
               Strg_TO_Chars(Strg:= CONCAT_STRING(IN1 := #TMP_strDef ,IN2 := DINT_TO_STRING(#INO_tDefects.tDefectsForReport.rgtDefects[#TMP_dIndexDef].dCoreWidth_um)),
                         pChars:=#TMP_dIndex,
                         Cnt=>#TMP_uiNumChar,
                         Chars:=#AUX_rgcDefectTelegram);
               #TMP_dIndex+=#TMP_uiNumChar;

               #AUX_rgcDefectTelegram[#TMP_dIndex] := #STRSEPARATOR;
               #TMP_dIndex+=1;

               //Defect distortion length
               #TMP_strDef := CONCAT_STRING(IN1 := #STRDEFECTDISTLENGTH ,IN2 := #TMP_strDefIndex);
               #TMP_strDef := CONCAT_STRING(IN1 := #TMP_strDef,IN2 := '=');

               Strg_TO_Chars(Strg:= CONCAT_STRING(IN1 := #TMP_strDef ,IN2 := DINT_TO_STRING(#INO_tDefects.tDefectsForReport.rgtDefects[#TMP_dIndexDef].dDistLength_um)),
                         pChars:=#TMP_dIndex,
                         Cnt=>#TMP_uiNumChar,
                         Chars:=#AUX_rgcDefectTelegram);
               #TMP_dIndex+=#TMP_uiNumChar;

               #AUX_rgcDefectTelegram[#TMP_dIndex] := #STRSEPARATOR;
               #TMP_dIndex+=1;

               //Defect distortion width
               #TMP_strDef := CONCAT_STRING(IN1 := #STRDEFECTDISTWIDTH ,IN2 := #TMP_strDefIndex);
               #TMP_strDef := CONCAT_STRING(IN1 := #TMP_strDef,IN2 := '=');

               Strg_TO_Chars(Strg:= CONCAT_STRING(IN1 := #TMP_strDef ,IN2 := DINT_TO_STRING(#INO_tDefects.tDefectsForReport.rgtDefects[#TMP_dIndexDef].dDistWidth_um)),
                         pChars:=#TMP_dIndex,
                         Cnt=>#TMP_uiNumChar,
                         Chars:=#AUX_rgcDefectTelegram);
               #TMP_dIndex+=#TMP_uiNumChar;

               #AUX_rgcDefectTelegram[#TMP_dIndex] := #STRSEPARATOR;
               #TMP_dIndex+=1;

               //Defect distortion optical value
               #TMP_strDef := CONCAT_STRING(IN1 := #STRDEFECTOPTVAL ,IN2 := #TMP_strDefIndex);
               #TMP_strDef := CONCAT_STRING(IN1 := #TMP_strDef,IN2 := '=');

               Strg_TO_Chars(Strg:= CONCAT_STRING(IN1 := #TMP_strDef ,IN2 := DINT_TO_STRING(#INO_tDefects.tDefectsForReport.rgtDefects[#TMP_dIndexDef].dOptValue_mdptr)),
                         pChars:=#TMP_dIndex,
                         Cnt=>#TMP_uiNumChar,
                         Chars:=#AUX_rgcDefectTelegram);
               #TMP_dIndex+=#TMP_uiNumChar;

               #AUX_rgcDefectTelegram[#TMP_dIndex] := #STRSEPARATOR;
               #TMP_dIndex+=1;

               //Defect string ID
               #TMP_strDef := CONCAT_STRING(IN1 := #STRDEFECTSCID ,IN2 := #TMP_strDefIndex);
               #TMP_strDef := CONCAT_STRING(IN1 := #TMP_strDef,IN2 := '=');

               Strg_TO_Chars(Strg:= CONCAT_STRING(IN1 := #TMP_strDef ,IN2 := #INO_tDefects.tDefectsForReport.rgtDefects[#TMP_dIndexDef].strDefectID),
                         pChars:=#TMP_dIndex,
                         Cnt=>#TMP_uiNumChar,
                         Chars:=#AUX_rgcDefectTelegram);
               #TMP_dIndex+=#TMP_uiNumChar;

               #AUX_rgcDefectTelegram[#TMP_dIndex] := #STRSEPARATOR;
               #TMP_dIndex+=1;

           END_FOR;

           //Compile the number of byte and set telegram available to  send
           #AUX_rgcDefectTelegram[#TMP_dIndex] := #STR_CR;
           #TMP_dIndex+=1;

           #AUX_rgcDefectTelegram[#TMP_dIndex] := #STR_LF;

           #AUX_dDefectTelegramNumByte := #TMP_dIndex + 1;

           IF #AUX_dDefectTelegramCounter >= #DMAXTELEGRAMCOUNTER THEN
               #AUX_dDefectTelegramCounter := 1;
           ELSE
               #AUX_dDefectTelegramCounter += 1;
           END_IF;

           #ST_xDefectTelegramAvail := TRUE;
           #INO_tDefects.tDefectsForReport.dNumberOfDefect := 0;

       END_IF;    

   END_IF;


   END_REGION BPS_DEFECTS_TELEGRAM

   REGION BPS_PLATE_TELEGRAM

   IF NOT #ST_xPlateTelegramAvail  AND #TMP_xSystemConnected  THEN

       //Search from the oldest one to send
       #TMP_dTail := #INO_tCaps.dTrackingTail;
       #TMP_xCapToSendFound := FALSE;

       WHILE (#TMP_dTail <> #INO_tCaps.dTrackingHead) DO

           IF (#INO_tCaps.rgtTrackCaps[#TMP_dTail].tCap.dID <> 0) AND 
                           ((#INO_tCaps.rgtTrackCaps[#TMP_dTail].tCap.tRequests.xUpdateDataBPSA AND #IN_xBPSServerA) OR 
                           (#INO_tCaps.rgtTrackCaps[#TMP_dTail].tCap.tRequests.xUpdateDataBPSB AND NOT #IN_xBPSServerA) (*OR #AUX_xResendAllPlate*))   THEN

               //New plate available to send. Copy the plate data on the local buffer and set the plate sent signal.
               #AUX_tCapToSend := #INO_tCaps.rgtTrackCaps[#TMP_dTail].tCap;
               IF #IN_xBPSServerA THEN
                   #INO_tCaps.rgtTrackCaps[#TMP_dTail].tCap.tRequests.xUpdateDataBPSA := FALSE;
               ELSE
                   #INO_tCaps.rgtTrackCaps[#TMP_dTail].tCap.tRequests.xUpdateDataBPSB := FALSE;
               END_IF;

               #TMP_xCapToSendFound := TRUE;

               EXIT;
           ELSE
               //Increment the tail
               IF (#TMP_dTail + 1) >= "DMAXTRACKCAP" THEN
                   #TMP_dTail := 0;
               ELSE
                   #TMP_dTail+= 1;
               END_IF;

           END_IF;
       END_WHILE;

       IF #TMP_xCapToSendFound THEN

           //Plate found start to prepare the respective telegram
           #TMP_dIndex := 0;

           #AUX_rgcPlateTelegram[#TMP_dIndex] := #STRPLATETELEGRAMID;
           #TMP_dIndex+=1;

           #AUX_rgcPlateTelegram[#TMP_dIndex] := #STRSEPARATOR;
           #TMP_dIndex+=1;

           Strg_TO_Chars(Strg:= CONCAT_STRING(IN1 := #STRPLATETELCOUNTER ,IN2 := DINT_TO_STRING(#AUX_dPlateTelegramCounter)),
                         pChars:=#TMP_dIndex,
                         Cnt=>#TMP_uiNumChar,
                         Chars:=#AUX_rgcPlateTelegram);
           #TMP_dIndex+=#TMP_uiNumChar;

           #AUX_rgcPlateTelegram[#TMP_dIndex] := #STRSEPARATOR;
           #TMP_dIndex+=1;

           Strg_TO_Chars(Strg:= CONCAT_STRING(IN1 := #STRCAPIDDESCR ,IN2 := DINT_TO_STRING(#AUX_tCapToSend.dID)),
                         pChars:=#TMP_dIndex,
                         Cnt=>#TMP_uiNumChar,
                         Chars:=#AUX_rgcPlateTelegram);
           #TMP_dIndex+=#TMP_uiNumChar;

           #AUX_rgcPlateTelegram[#TMP_dIndex] := #STRSEPARATOR;
           #TMP_dIndex+=1;

           Strg_TO_Chars(Strg:= CONCAT_STRING(IN1 := #STRCAPHEADPOS ,IN2 := DINT_TO_STRING(#AUX_tCapToSend.dHeadPositionBTC)),
                         pChars:=#TMP_dIndex,
                         Cnt=>#TMP_uiNumChar,
                         Chars:=#AUX_rgcPlateTelegram);
           #TMP_dIndex+=#TMP_uiNumChar;

           #AUX_rgcPlateTelegram[#TMP_dIndex] := #STRSEPARATOR;
           #TMP_dIndex+=1;

          Strg_TO_Chars(Strg:= CONCAT_STRING(IN1 := #STRCAPTAILPOS ,IN2 := DINT_TO_STRING(#AUX_tCapToSend.dTailPositionBTC)),
                         pChars:=#TMP_dIndex,
                         Cnt=>#TMP_uiNumChar,
                         Chars:=#AUX_rgcPlateTelegram);
           #TMP_dIndex+=#TMP_uiNumChar;

           #AUX_rgcPlateTelegram[#TMP_dIndex] := #STRSEPARATOR;
           #TMP_dIndex+=1;

          Strg_TO_Chars(Strg:= CONCAT_STRING(IN1 := #STRCAPLENGTH ,IN2 := DINT_TO_STRING(#AUX_tCapToSend.dLength_cmm)),
                         pChars:=#TMP_dIndex,
                         Cnt=>#TMP_uiNumChar,
                         Chars:=#AUX_rgcPlateTelegram);
           #TMP_dIndex+=#TMP_uiNumChar;

           #AUX_rgcPlateTelegram[#TMP_dIndex] := #STRSEPARATOR;
           #TMP_dIndex+=1;

          Strg_TO_Chars(Strg:= CONCAT_STRING(IN1 := #STRCAPWIDTH ,IN2 := DINT_TO_STRING(#AUX_tCapToSend.dWidth_cmm)),
                         pChars:=#TMP_dIndex,
                         Cnt=>#TMP_uiNumChar,
                         Chars:=#AUX_rgcPlateTelegram);
           #TMP_dIndex+=#TMP_uiNumChar;

           #AUX_rgcPlateTelegram[#TMP_dIndex] := #STRSEPARATOR;
           #TMP_dIndex+=1;

          Strg_TO_Chars(Strg:= CONCAT_STRING(IN1 := #STRCAPTHICK ,IN2 := DINT_TO_STRING(#AUX_tCapToSend.dThick_cmm)),
                         pChars:=#TMP_dIndex,
                         Cnt=>#TMP_uiNumChar,
                         Chars:=#AUX_rgcPlateTelegram);
           #TMP_dIndex+=#TMP_uiNumChar;

           #AUX_rgcPlateTelegram[#TMP_dIndex] := #STRSEPARATOR;
           #TMP_dIndex+=1;

           Strg_TO_Chars(Strg := CONCAT_STRING(IN1 := #STRCAPINDEX, IN2 := DINT_TO_STRING(#AUX_tCapToSend.dIndex)),
                         pChars := #TMP_dIndex,
                         Cnt => #TMP_uiNumChar,
                         Chars := #AUX_rgcPlateTelegram);
           #TMP_dIndex += #TMP_uiNumChar;

           #AUX_rgcPlateTelegram[#TMP_dIndex] := #STRSEPARATOR;
           #TMP_dIndex += 1;


          Strg_TO_Chars(Strg:= CONCAT_STRING(IN1 := #STRCAPFORMAT ,IN2 := DINT_TO_STRING(#AUX_tCapToSend.dFormat)),
                         pChars:=#TMP_dIndex,
                         Cnt=>#TMP_uiNumChar,
                         Chars:=#AUX_rgcPlateTelegram);
           #TMP_dIndex+=#TMP_uiNumChar;

           #AUX_rgcPlateTelegram[#TMP_dIndex] := #STRSEPARATOR;
           #TMP_dIndex+=1;

          Strg_TO_Chars(Strg:= CONCAT_STRING(IN1 := #STRCAPNUMLITE ,IN2 := DINT_TO_STRING(#AUX_tCapToSend.dNumLites)),
                         pChars:=#TMP_dIndex,
                         Cnt=>#TMP_uiNumChar,
                         Chars:=#AUX_rgcPlateTelegram);
           #TMP_dIndex+=#TMP_uiNumChar;

           #AUX_rgcPlateTelegram[#TMP_dIndex] := #STRSEPARATOR;
           #TMP_dIndex+=1;

          Strg_TO_Chars(Strg:= CONCAT_STRING(IN1 := #STRCAPREQGAP ,IN2 := DINT_TO_STRING(#AUX_tCapToSend.dReqGapForConv_cmm)),
                         pChars:=#TMP_dIndex,
                         Cnt=>#TMP_uiNumChar,
                         Chars:=#AUX_rgcPlateTelegram);
           #TMP_dIndex+=#TMP_uiNumChar;

           #AUX_rgcPlateTelegram[#TMP_dIndex] := #STRSEPARATOR;
           #TMP_dIndex+=1;

          Strg_TO_Chars(Strg:= CONCAT_STRING(IN1 := #STRCAPMAXCAP ,IN2 := DINT_TO_STRING(#AUX_tCapToSend.dMaxCapInConv)),
                         pChars:=#TMP_dIndex,
                         Cnt=>#TMP_uiNumChar,
                         Chars:=#AUX_rgcPlateTelegram);
           #TMP_dIndex+=#TMP_uiNumChar;

           #AUX_rgcPlateTelegram[#TMP_dIndex] := #STRSEPARATOR;
           #TMP_dIndex+=1;

          Strg_TO_Chars(Strg:= CONCAT_STRING(IN1 := #STRCAPCONVTOTLENGTH ,IN2 := DINT_TO_STRING(#AUX_tCapToSend.dConvTotLength_cmm)),
                         pChars:=#TMP_dIndex,
                         Cnt=>#TMP_uiNumChar,
                         Chars:=#AUX_rgcPlateTelegram);
           #TMP_dIndex+=#TMP_uiNumChar;

           #AUX_rgcPlateTelegram[#TMP_dIndex] := #STRSEPARATOR;
           #TMP_dIndex+=1;

          Strg_TO_Chars(Strg:= CONCAT_STRING(IN1 := #STRCAPGROSSWIDTH ,IN2 := DINT_TO_STRING(#AUX_tCapToSend.dGrossWidth_cmm)),
                         pChars:=#TMP_dIndex,
                         Cnt=>#TMP_uiNumChar,
                         Chars:=#AUX_rgcPlateTelegram);
           #TMP_dIndex+=#TMP_uiNumChar;

           #AUX_rgcPlateTelegram[#TMP_dIndex] := #STRSEPARATOR;
           #TMP_dIndex+=1;

          Strg_TO_Chars(Strg:= CONCAT_STRING(IN1 := #STRCAPNETWIDTH ,IN2 := DINT_TO_STRING(#AUX_tCapToSend.dNetWidth_cmm)),
                         pChars:=#TMP_dIndex,
                         Cnt=>#TMP_uiNumChar,
                         Chars:=#AUX_rgcPlateTelegram);
           #TMP_dIndex+=#TMP_uiNumChar;

           #AUX_rgcPlateTelegram[#TMP_dIndex] := #STRSEPARATOR;
           #TMP_dIndex+=1;

          Strg_TO_Chars(Strg:= CONCAT_STRING(IN1 := #STRCAPIDEDGEOPSIDE ,IN2 := DINT_TO_STRING(#AUX_tCapToSend.dDEdgeOpSide_cmm)),
                         pChars:=#TMP_dIndex,
                         Cnt=>#TMP_uiNumChar,
                         Chars:=#AUX_rgcPlateTelegram);
           #TMP_dIndex+=#TMP_uiNumChar;

           #AUX_rgcPlateTelegram[#TMP_dIndex] := #STRSEPARATOR;
           #TMP_dIndex+=1;

          Strg_TO_Chars(Strg:= CONCAT_STRING(IN1 := #STRCAPIDEDGEOPPOSIDE ,IN2 := DINT_TO_STRING(#AUX_tCapToSend.dDEdgeOppOpSide_cmm)),
                         pChars:=#TMP_dIndex,
                         Cnt=>#TMP_uiNumChar,
                         Chars:=#AUX_rgcPlateTelegram);
           #TMP_dIndex+=#TMP_uiNumChar;

           #AUX_rgcPlateTelegram[#TMP_dIndex] := #STRSEPARATOR;
           #TMP_dIndex+=1;

          Strg_TO_Chars(Strg:= CONCAT_STRING(IN1 := #STRCAPWANDER ,IN2 := DINT_TO_STRING(#AUX_tCapToSend.dEndCutWander_cmm)),
                         pChars:=#TMP_dIndex,
                         Cnt=>#TMP_uiNumChar,
                         Chars:=#AUX_rgcPlateTelegram);
           #TMP_dIndex+=#TMP_uiNumChar;

           #AUX_rgcPlateTelegram[#TMP_dIndex] := #STRSEPARATOR;
           #TMP_dIndex+=1;

          Strg_TO_Chars(Strg:= CONCAT_STRING(IN1 := #STRCAPNETWANDER ,IN2 := DINT_TO_STRING(#AUX_tCapToSend.dNetWander_cmm)),
                         pChars:=#TMP_dIndex,
                         Cnt=>#TMP_uiNumChar,
                         Chars:=#AUX_rgcPlateTelegram);
           #TMP_dIndex+=#TMP_uiNumChar;

           #AUX_rgcPlateTelegram[#TMP_dIndex] := #STRSEPARATOR;
           #TMP_dIndex+=1;

          Strg_TO_Chars(Strg:= CONCAT_STRING(IN1 := #STRCAPGROSSWANDER ,IN2 := DINT_TO_STRING(#AUX_tCapToSend.dGrossWander_cmm)),
                         pChars:=#TMP_dIndex,
                         Cnt=>#TMP_uiNumChar,
                         Chars:=#AUX_rgcPlateTelegram);
           #TMP_dIndex+=#TMP_uiNumChar;

           #AUX_rgcPlateTelegram[#TMP_dIndex] := #STRSEPARATOR;
           #TMP_dIndex+=1;

          Strg_TO_Chars(Strg:= CONCAT_STRING(IN1 := #STRCAPCOLOR ,IN2 := DINT_TO_STRING(#AUX_tCapToSend.dColor)),
                         pChars:=#TMP_dIndex,
                         Cnt=>#TMP_uiNumChar,
                         Chars:=#AUX_rgcPlateTelegram);
           #TMP_dIndex+=#TMP_uiNumChar;

           #AUX_rgcPlateTelegram[#TMP_dIndex] := #STRSEPARATOR;
           #TMP_dIndex+=1;

          Strg_TO_Chars(Strg:= CONCAT_STRING(IN1 := #STRCAPCOLORDESCR ,IN2 := #AUX_tCapToSend.strColorDescr),
                         pChars:=#TMP_dIndex,
                         Cnt=>#TMP_uiNumChar,
                         Chars:=#AUX_rgcPlateTelegram);
           #TMP_dIndex+=#TMP_uiNumChar;

           #AUX_rgcPlateTelegram[#TMP_dIndex] := #STRSEPARATOR;
           #TMP_dIndex+=1;

          Strg_TO_Chars(Strg:=CONCAT_STRING(IN1 := #STRCAPSYSMEAS ,IN2 := DINT_TO_STRING(#AUX_tCapToSend.dSystemMeasure)),
                         pChars:=#TMP_dIndex,
                         Cnt=>#TMP_uiNumChar,
                         Chars:=#AUX_rgcPlateTelegram);
           #TMP_dIndex+=#TMP_uiNumChar;

           #AUX_rgcPlateTelegram[#TMP_dIndex] := #STRSEPARATOR;
           #TMP_dIndex+=1;


           #TMP_dBridgeRequest := 0;
           #TMP_wBridgeMask := 0;

           IF #AUX_tCapToSend.tRequests.tYCutsData[0].xUseThisBridge THEN
               #TMP_dBridgeRequest := 1;
               GATHER(IN:=#AUX_tCapToSend.tRequests.tYCutsData[0].rgxHeadsRequest,
                                          OUT=>#TMP_wBridgeMask);

           ELSIF #AUX_tCapToSend.tRequests.tYCutsData[1].xUseThisBridge THEN
               #TMP_dBridgeRequest := 2;
               GATHER(IN:=#AUX_tCapToSend.tRequests.tYCutsData[1].rgxHeadsRequest,
                                          OUT=>#TMP_wBridgeMask);

           END_IF;

          Strg_TO_Chars(Strg:=CONCAT_STRING(IN1 := #STRCAPYCUTBRIDGESEL ,IN2 := DINT_TO_STRING(#TMP_dBridgeRequest)),
                         pChars:=#TMP_dIndex,
                         Cnt=>#TMP_uiNumChar,
                         Chars:=#AUX_rgcPlateTelegram);
           #TMP_dIndex+=#TMP_uiNumChar;

           #AUX_rgcPlateTelegram[#TMP_dIndex] := #STRSEPARATOR;
           #TMP_dIndex+=1;


          Strg_TO_Chars(Strg:=CONCAT_STRING(IN1 := #STRCAPYCUTHEADNUM ,IN2 := INT_TO_STRING(WORD_TO_INT(#TMP_wBridgeMask))),
                         pChars:=#TMP_dIndex,
                         Cnt=>#TMP_uiNumChar,
                         Chars:=#AUX_rgcPlateTelegram);
           #TMP_dIndex+=#TMP_uiNumChar;

           #AUX_rgcPlateTelegram[#TMP_dIndex] := #STRSEPARATOR;
           #TMP_dIndex+=1;



           FOR #TMP_dLiteIndex := 0 TO #AUX_tCapToSend.dNumLites - 1 DO

               #TMP_strFixLite := BYTE_TO_CHAR(CHAR_TO_BYTE(#STRLITEIDENT) + DINT_TO_BYTE(#TMP_dLiteIndex));

               #TMP_strTemp := CONCAT_STRING(IN1 := #TMP_strFixLite ,IN2 := #STRLITEID);

               Strg_TO_Chars(Strg:= CONCAT_STRING(IN1 := #TMP_strTemp ,IN2 := DINT_TO_STRING(#AUX_tCapToSend.rgtLites[#TMP_dLiteIndex].dID)),
                             pChars:=#TMP_dIndex,
                             Cnt=>#TMP_uiNumChar,
                             Chars:=#AUX_rgcPlateTelegram);
               #TMP_dIndex+=#TMP_uiNumChar;

               #AUX_rgcPlateTelegram[#TMP_dIndex] := #STRSEPARATOR;
               #TMP_dIndex+=1;

               #TMP_strTemp := CONCAT_STRING(IN1 := #TMP_strFixLite ,IN2 := #STRLITEPRODID);

               Strg_TO_Chars(Strg:= CONCAT_STRING(IN1 := #TMP_strTemp ,IN2 := DINT_TO_STRING(#AUX_tCapToSend.rgtLites[#TMP_dLiteIndex].dProductionID)),
                             pChars:=#TMP_dIndex,
                             Cnt=>#TMP_uiNumChar,
                             Chars:=#AUX_rgcPlateTelegram);
               #TMP_dIndex+=#TMP_uiNumChar;

               #AUX_rgcPlateTelegram[#TMP_dIndex] := #STRSEPARATOR;
               #TMP_dIndex+=1;

               #TMP_strTemp := CONCAT_STRING(IN1 := #TMP_strFixLite ,IN2 := #STRLITEPRODDESCR);

               Strg_TO_Chars(Strg:= CONCAT_STRING(IN1 := #TMP_strTemp ,IN2 :=#AUX_tCapToSend.rgtLites[#TMP_dLiteIndex].strProdDescr),
                             pChars:=#TMP_dIndex,
                             Cnt=>#TMP_uiNumChar,
                             Chars:=#AUX_rgcPlateTelegram);
               #TMP_dIndex+=#TMP_uiNumChar;

               #AUX_rgcPlateTelegram[#TMP_dIndex] := #STRSEPARATOR;
               #TMP_dIndex+=1;

               #TMP_strTemp := CONCAT_STRING(IN1 := #TMP_strFixLite ,IN2 := #STRLITEQUALID);

               Strg_TO_Chars(Strg:= CONCAT_STRING(IN1 := #TMP_strTemp ,IN2 := DINT_TO_STRING(#AUX_tCapToSend.rgtLites[#TMP_dLiteIndex].dQualityID)),
                             pChars:=#TMP_dIndex,
                             Cnt=>#TMP_uiNumChar,
                             Chars:=#AUX_rgcPlateTelegram);
               #TMP_dIndex+=#TMP_uiNumChar;

               #AUX_rgcPlateTelegram[#TMP_dIndex] := #STRSEPARATOR;
               #TMP_dIndex+=1;

               #TMP_strTemp := CONCAT_STRING(IN1 := #TMP_strFixLite ,IN2 := #STRLITEQUALDESCR);

               Strg_TO_Chars(Strg:= CONCAT_STRING(IN1 := #TMP_strTemp ,IN2 := #AUX_tCapToSend.rgtLites[#TMP_dLiteIndex].strQualityDescr),
                             pChars:=#TMP_dIndex,
                             Cnt=>#TMP_uiNumChar,
                             Chars:=#AUX_rgcPlateTelegram);
               #TMP_dIndex+=#TMP_uiNumChar;

               #AUX_rgcPlateTelegram[#TMP_dIndex] := #STRSEPARATOR;
               #TMP_dIndex+=1;

               #TMP_strTemp := CONCAT_STRING(IN1 := #TMP_strFixLite ,IN2 := #STRLITECAMERARECIPE);

               Strg_TO_Chars(Strg:= CONCAT_STRING(IN1 := #TMP_strTemp ,IN2 := DINT_TO_STRING(#AUX_tCapToSend.rgtLites[#TMP_dLiteIndex].dCameraRecipeID)),
                             pChars:=#TMP_dIndex,
                             Cnt=>#TMP_uiNumChar,
                             Chars:=#AUX_rgcPlateTelegram);
               #TMP_dIndex+=#TMP_uiNumChar;

               #AUX_rgcPlateTelegram[#TMP_dIndex] := #STRSEPARATOR;
               #TMP_dIndex+=1;

               #TMP_strTemp := CONCAT_STRING(IN1 := #TMP_strFixLite ,IN2 := #STRLITEWIDTH);

               Strg_TO_Chars(Strg:= CONCAT_STRING(IN1 := #TMP_strTemp ,IN2 := DINT_TO_STRING(#AUX_tCapToSend.rgtLites[#TMP_dLiteIndex].dWidth_cmm)),
                             pChars:=#TMP_dIndex,
                             Cnt=>#TMP_uiNumChar,
                             Chars:=#AUX_rgcPlateTelegram);
               #TMP_dIndex+=#TMP_uiNumChar;

               #AUX_rgcPlateTelegram[#TMP_dIndex] := #STRSEPARATOR;
               #TMP_dIndex+=1;

               #TMP_strTemp := CONCAT_STRING(IN1 := #TMP_strFixLite ,IN2 := #STRLITEBARYCENTRE);

               Strg_TO_Chars(Strg:= CONCAT_STRING(IN1 := #TMP_strTemp ,IN2 := DINT_TO_STRING(#AUX_tCapToSend.rgtLites[#TMP_dLiteIndex].dBarycentre_cmm)),
                             pChars:=#TMP_dIndex,
                             Cnt=>#TMP_uiNumChar,
                             Chars:=#AUX_rgcPlateTelegram);
               #TMP_dIndex+=#TMP_uiNumChar;

               #AUX_rgcPlateTelegram[#TMP_dIndex] := #STRSEPARATOR;
               #TMP_dIndex+=1;

               #TMP_strTemp := CONCAT_STRING(IN1 := #TMP_strFixLite ,IN2 := #STRLITECULLET);

               Strg_TO_Chars(Strg:= CONCAT_STRING(IN1 := #TMP_strTemp ,IN2 := DINT_TO_STRING(#AUX_tCapToSend.rgtLites[#TMP_dLiteIndex].dCulletCause)),
                             pChars:=#TMP_dIndex,
                             Cnt=>#TMP_uiNumChar,
                             Chars:=#AUX_rgcPlateTelegram);
               #TMP_dIndex+=#TMP_uiNumChar;

               #AUX_rgcPlateTelegram[#TMP_dIndex] := #STRSEPARATOR;
               #TMP_dIndex+=1;

               #TMP_strTemp := CONCAT_STRING(IN1 := #TMP_strFixLite ,IN2 := #STRLITEMAINDEST);

               Strg_TO_Chars(Strg:= CONCAT_STRING(IN1 := #TMP_strTemp ,IN2 := LINT_TO_STRING(#AUX_tCapToSend.rgtLites[#TMP_dLiteIndex].dMainDestination)),
                             pChars:=#TMP_dIndex,
                             Cnt=>#TMP_uiNumChar,
                             Chars:=#AUX_rgcPlateTelegram);
               #TMP_dIndex+=#TMP_uiNumChar;

               #AUX_rgcPlateTelegram[#TMP_dIndex] := #STRSEPARATOR;
               #TMP_dIndex+=1;

               #TMP_strTemp := CONCAT_STRING(IN1 := #TMP_strFixLite ,IN2 := #STRLITEALTDEST);

               Strg_TO_Chars(Strg:= CONCAT_STRING(IN1 := #TMP_strTemp ,IN2 := LINT_TO_STRING(#AUX_tCapToSend.rgtLites[#TMP_dLiteIndex].dAltDestination)),
                             pChars:=#TMP_dIndex,
                             Cnt=>#TMP_uiNumChar,
                             Chars:=#AUX_rgcPlateTelegram);
               #TMP_dIndex+=#TMP_uiNumChar;

               #AUX_rgcPlateTelegram[#TMP_dIndex] := #STRSEPARATOR;
               #TMP_dIndex+=1;

               #TMP_strTemp := CONCAT_STRING(IN1 := #TMP_strFixLite ,IN2 := #STRLITE2NDDEST);

               Strg_TO_Chars(Strg:= CONCAT_STRING(IN1 := #TMP_strTemp ,IN2 := LINT_TO_STRING(#AUX_tCapToSend.rgtLites[#TMP_dLiteIndex].d2ndDestionation)),
                             pChars:=#TMP_dIndex,
                             Cnt=>#TMP_uiNumChar,
                             Chars:=#AUX_rgcPlateTelegram);
               #TMP_dIndex+=#TMP_uiNumChar;

               #AUX_rgcPlateTelegram[#TMP_dIndex] := #STRSEPARATOR;
               #TMP_dIndex+=1;

              #TMP_strTemp := CONCAT_STRING(IN1 := #TMP_strFixLite ,IN2 := #STRLITESATPLATE);

               Strg_TO_Chars(Strg:= CONCAT_STRING(IN1 := #TMP_strTemp ,IN2 := DINT_TO_STRING(BOOL_TO_DINT(#AUX_tCapToSend.rgtLites[#TMP_dLiteIndex].xSaturationPlate))),
                             pChars:=#TMP_dIndex,
                             Cnt=>#TMP_uiNumChar,
                             Chars:=#AUX_rgcPlateTelegram);
               #TMP_dIndex+=#TMP_uiNumChar;

               #AUX_rgcPlateTelegram[#TMP_dIndex] := #STRSEPARATOR;
               #TMP_dIndex+=1;

           END_FOR; 

           //Compile the number of byte and set telegram available to  send
           #AUX_rgcPlateTelegram[#TMP_dIndex] := #STR_CR;
           #TMP_dIndex+=1;

           #AUX_rgcPlateTelegram[#TMP_dIndex] := #STR_LF;

           #AUX_dPlateTelegramNumByte := #TMP_dIndex + 1;

           IF #AUX_dPlateTelegramCounter >= #DMAXTELEGRAMCOUNTER THEN
               #AUX_dPlateTelegramCounter := 1;
           ELSE
               #AUX_dPlateTelegramCounter += 1;
           END_IF;

           #ST_xPlateTelegramAvail := TRUE;

       END_IF;
   END_IF;

   END_REGION BPS_PLATE_TELEGRAM

   REGION BPS_STATUS_TELEGRAM

   #AUX_dWaitingNextStatus_ms-= #INO_tInitialize.OUT_dExecutionTime_ms;

   IF #AUX_dWaitingNextStatus_ms < 0 THEN
       #AUX_dWaitingNextStatus_ms := 0;
   END_IF;

   //Prepare status telegram
   IF NOT #ST_xStatusTelegramAvail AND #AUX_dWaitingNextStatus_ms = 0  AND #TMP_xSystemConnected THEN

   //    #AUX_xResendAllStatus := TRUE;
       //Initialize waiting timer
       #AUX_dWaitingNextStatus_ms := #DDELAYSTATUSPACKET_MS;

       //Plate found start to prepare the respective telegram
       #TMP_dIndex := 0;

       #AUX_rgcStatusTelegram[#TMP_dIndex] := #STRSTATUSTELEGRAMID;
       #TMP_dIndex+=1;

       #AUX_rgcStatusTelegram[#TMP_dIndex] := #STRSEPARATOR;
       #TMP_dIndex+=1;

       Strg_TO_Chars(Strg:= CONCAT_STRING(IN1 := #STRSTATUSTELCOUNTER ,IN2 := DINT_TO_STRING(#AUX_dStatusTelegramCounter)),
                     pChars:=#TMP_dIndex,
                     Cnt=>#TMP_uiNumChar,
                     Chars:=#AUX_rgcStatusTelegram);
       #TMP_dIndex+=#TMP_uiNumChar;

       #AUX_rgcStatusTelegram[#TMP_dIndex] := #STRSEPARATOR;
       #TMP_dIndex+=1;

       Strg_TO_Chars(Strg:= CONCAT_STRING(IN1 := #STRSTATUSSERVCOUNTER ,IN2 := DINT_TO_STRING(#AUX_dStatusServerCounter)),
                     pChars:=#TMP_dIndex,
                     Cnt=>#TMP_uiNumChar,
                     Chars:=#AUX_rgcStatusTelegram);
       #TMP_dIndex+=#TMP_uiNumChar;

       #AUX_rgcStatusTelegram[#TMP_dIndex] := #STRSEPARATOR;
       #TMP_dIndex+=1;

       REGION BPS_STATUS_TELEGRAM_GENERAL

           IF ((#IN_tStatusGeneral.dActivePLC <> #AUX_tStatusGeneral.dActivePLC) OR #AUX_xResendAllStatus) THEN

               #AUX_tStatusGeneral.dActivePLC := #IN_tStatusGeneral.dActivePLC;

               Strg_TO_Chars(Strg := CONCAT_STRING(IN1 := #STRSTATUSACTIVEPLC, IN2 := DINT_TO_STRING(#AUX_tStatusGeneral.dActivePLC)),
                             pChars := #TMP_dIndex,
                             Cnt => #TMP_uiNumChar,
                             Chars := #AUX_rgcStatusTelegram);
               #TMP_dIndex += #TMP_uiNumChar;

               #AUX_rgcStatusTelegram[#TMP_dIndex] := #STRSEPARATOR;
               #TMP_dIndex += 1;

           END_IF;

           IF ((#IN_tStatusGeneral.dAutoRibSelection <> #AUX_tStatusGeneral.dAutoRibSelection) OR #AUX_xResendAllStatus) THEN

               #AUX_tStatusGeneral.dAutoRibSelection := #IN_tStatusGeneral.dAutoRibSelection;

               Strg_TO_Chars(Strg := CONCAT_STRING(IN1 := #STRSTATUSRIBSELEC, IN2 := DINT_TO_STRING(#AUX_tStatusGeneral.dAutoRibSelection)),
                             pChars := #TMP_dIndex,
                             Cnt => #TMP_uiNumChar,
                             Chars := #AUX_rgcStatusTelegram);
               #TMP_dIndex += #TMP_uiNumChar;

               #AUX_rgcStatusTelegram[#TMP_dIndex] := #STRSEPARATOR;
               #TMP_dIndex += 1;

           END_IF;

           IF ((#IN_tStatusGeneral.dExtOptSelected <> #AUX_tStatusGeneral.dExtOptSelected) OR #AUX_xResendAllStatus) THEN

               #AUX_tStatusGeneral.dExtOptSelected := #IN_tStatusGeneral.dExtOptSelected;

               Strg_TO_Chars(Strg := CONCAT_STRING(IN1 := #STRSTATUSEXTOPTSEL, IN2 := DINT_TO_STRING(#AUX_tStatusGeneral.dExtOptSelected)),
                             pChars := #TMP_dIndex,
                             Cnt => #TMP_uiNumChar,
                             Chars := #AUX_rgcStatusTelegram);
               #TMP_dIndex += #TMP_uiNumChar;

               #AUX_rgcStatusTelegram[#TMP_dIndex] := #STRSEPARATOR;
               #TMP_dIndex += 1;

           END_IF;

           IF ((#IN_tStatusGeneral.dOptimizerMode <> #AUX_tStatusGeneral.dOptimizerMode) OR #AUX_xResendAllStatus) THEN

               #AUX_tStatusGeneral.dOptimizerMode := #IN_tStatusGeneral.dOptimizerMode;

               Strg_TO_Chars(Strg := CONCAT_STRING(IN1 := #STRSTATUSOPTMODE, IN2 := DINT_TO_STRING(#AUX_tStatusGeneral.dOptimizerMode)),
                             pChars := #TMP_dIndex,
                             Cnt => #TMP_uiNumChar,
                             Chars := #AUX_rgcStatusTelegram);
               #TMP_dIndex += #TMP_uiNumChar;

               #AUX_rgcStatusTelegram[#TMP_dIndex] := #STRSEPARATOR;
               #TMP_dIndex += 1;

           END_IF;

           IF ((#IN_tStatusGeneral.dOptStatus <> #AUX_tStatusGeneral.dOptStatus) OR #AUX_xResendAllStatus) THEN

               #AUX_tStatusGeneral.dOptStatus := #IN_tStatusGeneral.dOptStatus;

               Strg_TO_Chars(Strg := CONCAT_STRING(IN1 := #STRSTATUSOPTSTATUS, IN2 := DINT_TO_STRING(#AUX_tStatusGeneral.dOptStatus)),
                             pChars := #TMP_dIndex,
                             Cnt => #TMP_uiNumChar,
                             Chars := #AUX_rgcStatusTelegram);
               #TMP_dIndex += #TMP_uiNumChar;

               #AUX_rgcStatusTelegram[#TMP_dIndex] := #STRSEPARATOR;
               #TMP_dIndex += 1;

           END_IF;

           IF ((#IN_tStatusGeneral.dRibbonModality <> #AUX_tStatusGeneral.dRibbonModality) OR #AUX_xResendAllStatus) THEN

               #AUX_tStatusGeneral.dRibbonModality := #IN_tStatusGeneral.dRibbonModality;

               Strg_TO_Chars(Strg := CONCAT_STRING(IN1 := #STRSTATUSRIBMODE, IN2 := DINT_TO_STRING(#AUX_tStatusGeneral.dRibbonModality)),
                             pChars := #TMP_dIndex,
                             Cnt => #TMP_uiNumChar,
                             Chars := #AUX_rgcStatusTelegram);
               #TMP_dIndex += #TMP_uiNumChar;

               #AUX_rgcStatusTelegram[#TMP_dIndex] := #STRSEPARATOR;
               #TMP_dIndex += 1;

           END_IF;

           IF ((#IN_tStatusGeneral.dScanStatus <> #AUX_tStatusGeneral.dScanStatus) OR #AUX_xResendAllStatus) THEN

               #AUX_tStatusGeneral.dScanStatus := #IN_tStatusGeneral.dScanStatus;

               Strg_TO_Chars(Strg := CONCAT_STRING(IN1 := #STRSTATUSSCANNERSTATUS, IN2 := DINT_TO_STRING(#AUX_tStatusGeneral.dScanStatus)),
                             pChars := #TMP_dIndex,
                             Cnt => #TMP_uiNumChar,
                             Chars := #AUX_rgcStatusTelegram);
               #TMP_dIndex += #TMP_uiNumChar;

               #AUX_rgcStatusTelegram[#TMP_dIndex] := #STRSEPARATOR;
               #TMP_dIndex += 1;

           END_IF;

           IF ((#IN_tStatusGeneral.dTypeWanderSel <> #AUX_tStatusGeneral.dTypeWanderSel) OR #AUX_xResendAllStatus) THEN

               #AUX_tStatusGeneral.dTypeWanderSel := #IN_tStatusGeneral.dTypeWanderSel;

               Strg_TO_Chars(Strg := CONCAT_STRING(IN1 := #STRSTATUSTYPEWANDER, IN2 := DINT_TO_STRING(#AUX_tStatusGeneral.dTypeWanderSel)),
                             pChars := #TMP_dIndex,
                             Cnt => #TMP_uiNumChar,
                             Chars := #AUX_rgcStatusTelegram);
               #TMP_dIndex += #TMP_uiNumChar;

               #AUX_rgcStatusTelegram[#TMP_dIndex] := #STRSEPARATOR;
               #TMP_dIndex += 1;

           END_IF;

           IF ((#IN_tStatusGeneral.dScanGrossWidth_cmm <> #AUX_tStatusGeneral.dScanGrossWidth_cmm) OR #AUX_xResendAllStatus) THEN

               #AUX_tStatusGeneral.dScanGrossWidth_cmm := #IN_tStatusGeneral.dScanGrossWidth_cmm;

               Strg_TO_Chars(Strg := CONCAT_STRING(IN1 := #STRSTATUSSCANNERGROSSWIDTH, IN2 := DINT_TO_STRING(#AUX_tStatusGeneral.dScanGrossWidth_cmm)),
                             pChars := #TMP_dIndex,
                             Cnt => #TMP_uiNumChar,
                             Chars := #AUX_rgcStatusTelegram);
               #TMP_dIndex += #TMP_uiNumChar;

               #AUX_rgcStatusTelegram[#TMP_dIndex] := #STRSEPARATOR;
               #TMP_dIndex += 1;

           END_IF;

           IF ((#IN_tStatusGeneral.dScanNetWidth_cmm <> #AUX_tStatusGeneral.dScanNetWidth_cmm) OR #AUX_xResendAllStatus) THEN

               #AUX_tStatusGeneral.dScanNetWidth_cmm := #IN_tStatusGeneral.dScanNetWidth_cmm;

               Strg_TO_Chars(Strg := CONCAT_STRING(IN1 := #STRSTATUSSCANNERNETWIDTH, IN2 := DINT_TO_STRING(#AUX_tStatusGeneral.dScanNetWidth_cmm)),
                             pChars := #TMP_dIndex,
                             Cnt => #TMP_uiNumChar,
                             Chars := #AUX_rgcStatusTelegram);
               #TMP_dIndex += #TMP_uiNumChar;

               #AUX_rgcStatusTelegram[#TMP_dIndex] := #STRSEPARATOR;
               #TMP_dIndex += 1;

           END_IF;

           IF ((#IN_tStatusGeneral.dScanGrossWander_cmm <> #AUX_tStatusGeneral.dScanGrossWander_cmm) OR #AUX_xResendAllStatus) THEN

               #AUX_tStatusGeneral.dScanGrossWander_cmm := #IN_tStatusGeneral.dScanGrossWander_cmm;

               Strg_TO_Chars(Strg := CONCAT_STRING(IN1 := #STRSTATUSSCANNERGROSSWANDER, IN2 := DINT_TO_STRING(#AUX_tStatusGeneral.dScanGrossWander_cmm)),
                             pChars := #TMP_dIndex,
                             Cnt => #TMP_uiNumChar,
                             Chars := #AUX_rgcStatusTelegram);
               #TMP_dIndex += #TMP_uiNumChar;

               #AUX_rgcStatusTelegram[#TMP_dIndex] := #STRSEPARATOR;
               #TMP_dIndex += 1;

           END_IF;

           IF ((#IN_tStatusGeneral.dScanNetWander_cmm <> #AUX_tStatusGeneral.dScanNetWander_cmm) OR #AUX_xResendAllStatus) THEN

               #AUX_tStatusGeneral.dScanNetWander_cmm := #IN_tStatusGeneral.dScanNetWander_cmm;

               Strg_TO_Chars(Strg := CONCAT_STRING(IN1 := #STRSTATUSSCANNERNETWANDER, IN2 := DINT_TO_STRING(#AUX_tStatusGeneral.dScanNetWander_cmm)),
                             pChars := #TMP_dIndex,
                             Cnt => #TMP_uiNumChar,
                             Chars := #AUX_rgcStatusTelegram);
               #TMP_dIndex += #TMP_uiNumChar;

               #AUX_rgcStatusTelegram[#TMP_dIndex] := #STRSEPARATOR;
               #TMP_dIndex += 1;

           END_IF;

           IF ((#IN_tStatusGeneral.dWanderRecoveryThr_cmm <> #AUX_tStatusGeneral.dWanderRecoveryThr_cmm) OR #AUX_xResendAllStatus) THEN

               #AUX_tStatusGeneral.dWanderRecoveryThr_cmm := #IN_tStatusGeneral.dWanderRecoveryThr_cmm;

               Strg_TO_Chars(Strg := CONCAT_STRING(IN1 := #STRSTATUSWANDRECTHR, IN2 := DINT_TO_STRING(#AUX_tStatusGeneral.dWanderRecoveryThr_cmm)),
                             pChars := #TMP_dIndex,
                             Cnt => #TMP_uiNumChar,
                             Chars := #AUX_rgcStatusTelegram);
               #TMP_dIndex += #TMP_uiNumChar;

               #AUX_rgcStatusTelegram[#TMP_dIndex] := #STRSEPARATOR;
               #TMP_dIndex += 1;

           END_IF;

           IF ((#IN_tStatusGeneral.dYC1WandRec_cmm <> #AUX_tStatusGeneral.dYC1WandRec_cmm) OR #AUX_xResendAllStatus) THEN

               #AUX_tStatusGeneral.dYC1WandRec_cmm := #IN_tStatusGeneral.dYC1WandRec_cmm;

               Strg_TO_Chars(Strg := CONCAT_STRING(IN1 := #STRSTATUSWANDYC1, IN2 := DINT_TO_STRING(#AUX_tStatusGeneral.dYC1WandRec_cmm)),
                             pChars := #TMP_dIndex,
                             Cnt => #TMP_uiNumChar,
                             Chars := #AUX_rgcStatusTelegram);
               #TMP_dIndex += #TMP_uiNumChar;

               #AUX_rgcStatusTelegram[#TMP_dIndex] := #STRSEPARATOR;
               #TMP_dIndex += 1;

           END_IF;

           IF ((#IN_tStatusGeneral.dYC2WandRec_cmm <> #AUX_tStatusGeneral.dYC2WandRec_cmm) OR #AUX_xResendAllStatus) THEN

               #AUX_tStatusGeneral.dYC2WandRec_cmm := #IN_tStatusGeneral.dYC2WandRec_cmm;

               Strg_TO_Chars(Strg := CONCAT_STRING(IN1 := #STRSTATUSWANDYC2, IN2 := DINT_TO_STRING(#AUX_tStatusGeneral.dYC2WandRec_cmm)),
                             pChars := #TMP_dIndex,
                             Cnt => #TMP_uiNumChar,
                             Chars := #AUX_rgcStatusTelegram);
               #TMP_dIndex += #TMP_uiNumChar;

               #AUX_rgcStatusTelegram[#TMP_dIndex] := #STRSEPARATOR;
               #TMP_dIndex += 1;

           END_IF;

       END_REGION

       REGION BPS_STATUS_TELEGRAM_ENCODER


       //Encoder statuses

       #AUX_tStatusEncoder.dActualBTC_cmm := #IN_tStatusEncoder.dActualBTC_cmm;        

       Strg_TO_Chars(Strg:= CONCAT_STRING(IN1 := #STRSTATUSBTC ,IN2 := DINT_TO_STRING(#IN_tStatusEncoder.dActualBTC_cmm)),
                     pChars:=#TMP_dIndex,
                     Cnt=>#TMP_uiNumChar,
                     Chars:=#AUX_rgcStatusTelegram);
       #TMP_dIndex+=#TMP_uiNumChar;

       #AUX_rgcStatusTelegram[#TMP_dIndex] := #STRSEPARATOR;
       #TMP_dIndex+=1;

       IF (#IN_tStatusEncoder.dTrackSpeed_mm_min <> #AUX_tStatusEncoder.dTrackSpeed_mm_min) OR (#AUX_xResendAllStatus) THEN

           #AUX_tStatusEncoder.dTrackSpeed_mm_min := #IN_tStatusEncoder.dTrackSpeed_mm_min;

           Strg_TO_Chars(Strg := CONCAT_STRING(IN1 := #STRSTATUSLEHRSPEED, IN2 := DINT_TO_STRING(#IN_tStatusEncoder.dTrackSpeed_mm_min)),
                         pChars := #TMP_dIndex,
                         Cnt => #TMP_uiNumChar,
                         Chars := #AUX_rgcStatusTelegram);
           #TMP_dIndex += #TMP_uiNumChar;

           #AUX_rgcStatusTelegram[#TMP_dIndex] := #STRSEPARATOR;
           #TMP_dIndex += 1;

       END_IF;

       IF (#IN_dLineSpeed_mm_min <> #AUX_dLineSpeed_mm_min) OR (#AUX_xResendAllStatus) THEN

           #AUX_dLineSpeed_mm_min := #IN_dLineSpeed_mm_min;

           Strg_TO_Chars(Strg:= CONCAT_STRING(IN1 := #STRSTATUSTRACKSPEED ,IN2 := DINT_TO_STRING(#IN_dLineSpeed_mm_min)),
                         pChars:=#TMP_dIndex,
                         Cnt=>#TMP_uiNumChar,
                         Chars:=#AUX_rgcStatusTelegram);
           #TMP_dIndex+=#TMP_uiNumChar;

           #AUX_rgcStatusTelegram[#TMP_dIndex] := #STRSEPARATOR;
           #TMP_dIndex+=1;

       END_IF;

       IF (#IN_tStatusEncoder.dActSelEnc <> #AUX_tStatusEncoder.dActSelEnc) OR (#AUX_xResendAllStatus) THEN

           #AUX_tStatusEncoder.dActSelEnc := #IN_tStatusEncoder.dActSelEnc;        

           Strg_TO_Chars(Strg:= CONCAT_STRING(IN1 := #STRSTATUSACTSELENC ,IN2 := DINT_TO_STRING(#IN_tStatusEncoder.dActSelEnc)),
                         pChars:=#TMP_dIndex,
                         Cnt=>#TMP_uiNumChar,
                         Chars:=#AUX_rgcStatusTelegram);
           #TMP_dIndex+=#TMP_uiNumChar;

           #AUX_rgcStatusTelegram[#TMP_dIndex] := #STRSEPARATOR;
           #TMP_dIndex+=1;

       END_IF;

       END_REGION BPS_STATUS_TELEGRAM_ENCODER

       REGION BPS_STATUS_TELEGRAM_DIGITIZER1

       //Digitizer 1 status
       IF (#IN_tStatusDigitizer_1.dActualEncoderSpeed_mm_min <> #AUX_tStatusDigitizer_1.dActualEncoderSpeed_mm_min) OR (#AUX_xResendAllStatus) THEN

           #AUX_tStatusDigitizer_1.dActualEncoderSpeed_mm_min := #IN_tStatusDigitizer_1.dActualEncoderSpeed_mm_min;        

           Strg_TO_Chars(Strg:= CONCAT_STRING(IN1 := #STRSTATUSDGT1SPEED ,IN2 := DINT_TO_STRING(#IN_tStatusDigitizer_1.dActualEncoderSpeed_mm_min)),
                         pChars:=#TMP_dIndex,
                         Cnt=>#TMP_uiNumChar,
                         Chars:=#AUX_rgcStatusTelegram);
           #TMP_dIndex+=#TMP_uiNumChar;

           #AUX_rgcStatusTelegram[#TMP_dIndex] := #STRSEPARATOR;
           #TMP_dIndex+=1;

       END_IF;

       IF (#IN_tStatusDigitizer_1.dEncoderStatus <> #AUX_tStatusDigitizer_1.dEncoderStatus) OR (#AUX_xResendAllStatus) THEN

           #AUX_tStatusDigitizer_1.dEncoderStatus := #IN_tStatusDigitizer_1.dEncoderStatus;        

           Strg_TO_Chars(Strg:= CONCAT_STRING(IN1 := #STRSTATUSDGT1STATUS ,IN2 := DINT_TO_STRING(#IN_tStatusDigitizer_1.dEncoderStatus)),
                         pChars:=#TMP_dIndex,
                         Cnt=>#TMP_uiNumChar,
                         Chars:=#AUX_rgcStatusTelegram);
           #TMP_dIndex+=#TMP_uiNumChar;

           #AUX_rgcStatusTelegram[#TMP_dIndex] := #STRSEPARATOR;
           #TMP_dIndex+=1;

       END_IF;

       IF (#IN_tStatusDigitizer_1.dDistanceSnapRoll_cmm <> #AUX_tStatusDigitizer_1.dDistanceSnapRoll_cmm) OR (#AUX_xResendAllStatus) THEN

           #AUX_tStatusDigitizer_1.dDistanceSnapRoll_cmm := #IN_tStatusDigitizer_1.dDistanceSnapRoll_cmm;        

           Strg_TO_Chars(Strg:= CONCAT_STRING(IN1 := #STRSTATUSDGT1DISTSNAP ,IN2 := DINT_TO_STRING(#IN_tStatusDigitizer_1.dDistanceSnapRoll_cmm)),
                         pChars:=#TMP_dIndex,
                         Cnt=>#TMP_uiNumChar,
                         Chars:=#AUX_rgcStatusTelegram);
           #TMP_dIndex+=#TMP_uiNumChar;

           #AUX_rgcStatusTelegram[#TMP_dIndex] := #STRSEPARATOR;
           #TMP_dIndex+=1;

       END_IF;

       END_REGION BPS_STATUS_TELEGRAM_DIGITIZER1

       REGION BPS_STATUS_TELEGRAM_DIGITIZER2

       //Digitizer 2 status
       IF (#IN_tStatusDigitizer_2.dActualEncoderSpeed_mm_min <> #AUX_tStatusDigitizer_2.dActualEncoderSpeed_mm_min) OR (#AUX_xResendAllStatus) THEN

           #AUX_tStatusDigitizer_2.dActualEncoderSpeed_mm_min := #IN_tStatusDigitizer_2.dActualEncoderSpeed_mm_min;        

           Strg_TO_Chars(Strg:= CONCAT_STRING(IN1 := #STRSTATUSDGT2SPEED ,IN2 := DINT_TO_STRING(#IN_tStatusDigitizer_2.dActualEncoderSpeed_mm_min)),
                         pChars:=#TMP_dIndex,
                         Cnt=>#TMP_uiNumChar,
                         Chars:=#AUX_rgcStatusTelegram);
           #TMP_dIndex+=#TMP_uiNumChar;

           #AUX_rgcStatusTelegram[#TMP_dIndex] := #STRSEPARATOR;
           #TMP_dIndex+=1;

       END_IF;

       IF (#IN_tStatusDigitizer_2.dEncoderStatus <> #AUX_tStatusDigitizer_2.dEncoderStatus) OR (#AUX_xResendAllStatus) THEN

           #AUX_tStatusDigitizer_2.dEncoderStatus := #IN_tStatusDigitizer_2.dEncoderStatus;        

           Strg_TO_Chars(Strg:= CONCAT_STRING(IN1 := #STRSTATUSDGT2STATUS ,IN2 := DINT_TO_STRING(#IN_tStatusDigitizer_2.dEncoderStatus)),
                         pChars:=#TMP_dIndex,
                         Cnt=>#TMP_uiNumChar,
                         Chars:=#AUX_rgcStatusTelegram);
           #TMP_dIndex+=#TMP_uiNumChar;

           #AUX_rgcStatusTelegram[#TMP_dIndex] := #STRSEPARATOR;
           #TMP_dIndex+=1;

       END_IF;

       IF (#IN_tStatusDigitizer_2.dDistanceSnapRoll_cmm <> #AUX_tStatusDigitizer_2.dDistanceSnapRoll_cmm) OR (#AUX_xResendAllStatus) THEN

           #AUX_tStatusDigitizer_2.dDistanceSnapRoll_cmm := #IN_tStatusDigitizer_2.dDistanceSnapRoll_cmm;        

           Strg_TO_Chars(Strg:= CONCAT_STRING(IN1 := #STRSTATUSDGT2DISTSNAP ,IN2 := DINT_TO_STRING(#IN_tStatusDigitizer_2.dDistanceSnapRoll_cmm)),
                         pChars:=#TMP_dIndex,
                         Cnt=>#TMP_uiNumChar,
                         Chars:=#AUX_rgcStatusTelegram);
           #TMP_dIndex+=#TMP_uiNumChar;

           #AUX_rgcStatusTelegram[#TMP_dIndex] := #STRSEPARATOR;
           #TMP_dIndex+=1;

       END_IF;

       END_REGION BPS_STATUS_TELEGRAM_DIGITIZER2

       REGION BPS_STATUS_TELEGRAM_XCUTS

       FOR #TMP_dXCutIndex := 0 TO "DMAXXHEADS_IND" DO

           #TMP_strXCutIndex := DINT_TO_STRING(#TMP_dXCutIndex + 1);   

           #TMP_strXCutIndex := DELETE(IN:=#TMP_strXCutIndex, L:=1, P:=1);

           IF (#IN_rgtStatusXCuts[#TMP_dXCutIndex].dActualCarriagePos_cmm <> #AUX_rgtStatusXCuts[#TMP_dXCutIndex].dActualCarriagePos_cmm) OR (#AUX_xResendAllStatus) THEN

               #AUX_rgtStatusXCuts[#TMP_dXCutIndex].dActualCarriagePos_cmm := #IN_rgtStatusXCuts[#TMP_dXCutIndex].dActualCarriagePos_cmm;        

               #TMP_strTemp := CONCAT_STRING(IN1 := #STRSTATUSXCUTACTPOS ,IN2 := #TMP_strXCutIndex);
               #TMP_strTemp := CONCAT_STRING(IN1 := #TMP_strTemp ,IN2 := '=');

               Strg_TO_Chars(Strg:= CONCAT_STRING(IN1 := #TMP_strTemp ,IN2 := DINT_TO_STRING(#IN_rgtStatusXCuts[#TMP_dXCutIndex].dActualCarriagePos_cmm)),
                         pChars:=#TMP_dIndex,
                         Cnt=>#TMP_uiNumChar,
                         Chars:=#AUX_rgcStatusTelegram);
               #TMP_dIndex+=#TMP_uiNumChar;

               #AUX_rgcStatusTelegram[#TMP_dIndex] := #STRSEPARATOR;
               #TMP_dIndex+=1;
           END_IF;

           IF (#IN_rgtStatusXCuts[#TMP_dXCutIndex].dDistanceFromSnaproll_cmm <> #AUX_rgtStatusXCuts[#TMP_dXCutIndex].dDistanceFromSnaproll_cmm) OR (#AUX_xResendAllStatus) THEN

               #AUX_rgtStatusXCuts[#TMP_dXCutIndex].dDistanceFromSnaproll_cmm := #IN_rgtStatusXCuts[#TMP_dXCutIndex].dDistanceFromSnaproll_cmm;        

               #TMP_strTemp := CONCAT_STRING(IN1 := #STRSTATUSXCUTDISTSNAP ,IN2 := #TMP_strXCutIndex);
               #TMP_strTemp := CONCAT_STRING(IN1 := #TMP_strTemp ,IN2 := '=');

               Strg_TO_Chars(Strg:= CONCAT_STRING(IN1 := #TMP_strTemp ,IN2 := DINT_TO_STRING(#IN_rgtStatusXCuts[#TMP_dXCutIndex].dDistanceFromSnaproll_cmm)),
                         pChars:=#TMP_dIndex,
                         Cnt=>#TMP_uiNumChar,
                         Chars:=#AUX_rgcStatusTelegram);
               #TMP_dIndex+=#TMP_uiNumChar;

               #AUX_rgcStatusTelegram[#TMP_dIndex] := #STRSEPARATOR;
               #TMP_dIndex+=1;
           END_IF;

           IF (#IN_rgtStatusXCuts[#TMP_dXCutIndex].dStatus <> #AUX_rgtStatusXCuts[#TMP_dXCutIndex].dStatus) OR (#AUX_xResendAllStatus) THEN

               #AUX_rgtStatusXCuts[#TMP_dXCutIndex].dStatus := #IN_rgtStatusXCuts[#TMP_dXCutIndex].dStatus;        

               #TMP_strTemp := CONCAT_STRING(IN1 := #STRSTATUSXCUTSTATUS ,IN2 := #TMP_strXCutIndex);
               #TMP_strTemp := CONCAT_STRING(IN1 := #TMP_strTemp ,IN2 := '=');

               Strg_TO_Chars(Strg:= CONCAT_STRING(IN1 := #TMP_strTemp ,IN2 := DINT_TO_STRING(#IN_rgtStatusXCuts[#TMP_dXCutIndex].dStatus)),
                         pChars:=#TMP_dIndex,
                         Cnt=>#TMP_uiNumChar,
                         Chars:=#AUX_rgcStatusTelegram);
               #TMP_dIndex+=#TMP_uiNumChar;

               #AUX_rgcStatusTelegram[#TMP_dIndex] := #STRSEPARATOR;
               #TMP_dIndex+=1;
           END_IF;

           IF (#IN_rgtStatusXCuts[#TMP_dXCutIndex].dXCutActualStatus <> #AUX_rgtStatusXCuts[#TMP_dXCutIndex].dXCutActualStatus) OR (#AUX_xResendAllStatus) THEN

               #AUX_rgtStatusXCuts[#TMP_dXCutIndex].dXCutActualStatus := #IN_rgtStatusXCuts[#TMP_dXCutIndex].dXCutActualStatus;        

               #TMP_strTemp := CONCAT_STRING(IN1 := #STRSTATUSXCUTACTSTATUS ,IN2 := #TMP_strXCutIndex);
               #TMP_strTemp := CONCAT_STRING(IN1 := #TMP_strTemp ,IN2 := '=');

               Strg_TO_Chars(Strg:= CONCAT_STRING(IN1 := #TMP_strTemp ,IN2 := DINT_TO_STRING(#IN_rgtStatusXCuts[#TMP_dXCutIndex].dXCutActualStatus)),
                         pChars:=#TMP_dIndex,
                         Cnt=>#TMP_uiNumChar,
                         Chars:=#AUX_rgcStatusTelegram);
               #TMP_dIndex+=#TMP_uiNumChar;

               #AUX_rgcStatusTelegram[#TMP_dIndex] := #STRSEPARATOR;
               #TMP_dIndex+=1;
           END_IF;

       END_FOR;

       END_REGION BPS_STATUS_TELEGRAM_XCUTS

       REGION BPS_STATUS_TELEGRAM_MARKERS

       FOR #TMP_dMarkerIndex := 0  TO "DMAXMARKERS_IND" DO

           #TMP_strMarkerIndex := DINT_TO_STRING(#TMP_dMarkerIndex + 1);

           #TMP_strMarkerIndex := DELETE(IN:= #TMP_strMarkerIndex, L:=1,P:=1);

           IF (#IN_rgtStatusMarkers[#TMP_dMarkerIndex].dActualCarriagePos_cmm <> #AUX_rgtStatusMarkers[#TMP_dMarkerIndex].dActualCarriagePos_cmm) OR (#AUX_xResendAllStatus) OR TRUE THEN

               #AUX_rgtStatusMarkers[#TMP_dMarkerIndex].dActualCarriagePos_cmm := #IN_rgtStatusMarkers[#TMP_dMarkerIndex].dActualCarriagePos_cmm;        

               #TMP_strTemp := CONCAT_STRING(IN1 := #STRSTATUSMARKACTPOS ,IN2 := #TMP_strMarkerIndex);
               #TMP_strTemp := CONCAT_STRING(IN1 := #TMP_strTemp ,IN2 := '=');

               Strg_TO_Chars(Strg:= CONCAT_STRING(IN1 := #TMP_strTemp ,IN2 := DINT_TO_STRING(#IN_rgtStatusMarkers[#TMP_dMarkerIndex].dActualCarriagePos_cmm)),
                         pChars:=#TMP_dIndex,
                         Cnt=>#TMP_uiNumChar,
                         Chars:=#AUX_rgcStatusTelegram);
               #TMP_dIndex+=#TMP_uiNumChar;

               #AUX_rgcStatusTelegram[#TMP_dIndex] := #STRSEPARATOR;
               #TMP_dIndex+=1;
           END_IF;



    (*       IF (#IN_rgtStatusMarkers[#TMP_dMarkerIndex].dDistanceFromSnaproll_cmm <> #AUX_rgtStatusMarkers[#TMP_dMarkerIndex].dDistanceFromSnaproll_cmm) OR (#AUX_xResendAllStatus) THEN

               #AUX_rgtStatusMarkers[#TMP_dMarkerIndex].dDistanceFromSnaproll_cmm := #IN_rgtStatusMarkers[#TMP_dMarkerIndex].dDistanceFromSnaproll_cmm;        

               #TMP_strTemp := CONCAT_STRING(IN1 := #STRSTATUSMARKDISTSNAP ,IN2 := #TMP_strMarkerIndex);
               #TMP_strTemp := CONCAT_STRING(IN1 := #TMP_strTemp ,IN2 := '=');

               Strg_TO_Chars(Strg:= CONCAT_STRING(IN1 := #TMP_strTemp ,IN2 := DINT_TO_STRING(#IN_rgtStatusMarkers[#TMP_dMarkerIndex].dDistanceFromSnaproll_cmm)),
                         pChars:=#TMP_dIndex,
                         Cnt=>#TMP_uiNumChar,
                         Chars:=#AUX_rgcStatusTelegram);
               #TMP_dIndex+=#TMP_uiNumChar;

               #AUX_rgcStatusTelegram[#TMP_dIndex] := #STRSEPARATOR;
               #TMP_dIndex+=1;
           END_IF;

           IF (#IN_rgtStatusMarkers[#TMP_dMarkerIndex].dStatus <> #AUX_rgtStatusMarkers[#TMP_dMarkerIndex].dStatus) OR (#AUX_xResendAllStatus) THEN

               #AUX_rgtStatusMarkers[#TMP_dMarkerIndex].dStatus := #IN_rgtStatusMarkers[#TMP_dMarkerIndex].dStatus;        

               #TMP_strTemp := CONCAT_STRING(IN1 := #STRSTATUSMARKSTATUS ,IN2 := #TMP_strMarkerIndex);
               #TMP_strTemp := CONCAT_STRING(IN1 := #TMP_strTemp ,IN2 := '=');

